
                       #INO_FB_Markers(IN_tNewMissionData := #TMP_tNewMisMark,
                                             IN_xStandardFBCall := FALSE,
                                             INO_xCallAddTank := #TMP_xCallAddTank,
                                             INO_tEnc := "DB_Encoder",INO_tRibbon := "DB_RibbonData");

                   END_IF;
               END_FOR;
           END_IF;
       END_IF;
   END_IF;

   //Manage received big telegram
   IF #FB_TRecvBig.DONE THEN

       //Check the packet telegram
       #TMP_dSerializePos := 0;
       #TMP_iReturn := Deserialize(SRC_ARRAY:=#AUX_rgb1000RecvBytePck, DEST_VARIABLE=>#TMP_dValue, POS:=#TMP_dSerializePos);

       IF #TMP_dValue = #DPLATEPACKTIDENT THEN

           #TMP_dSerializePos := 0;
           #TMP_iReturn := Deserialize(SRC_ARRAY:=#AUX_rgb1000RecvBytePck, DEST_VARIABLE=>#AUX_tPlatePacket, POS:=#TMP_dSerializePos);

           //Copy the plate to the buffer
           IF #AUX_dNumPlatePacket < #DMAXPLATEPACKET THEN

               #AUX_rgtPlatePacketArray[#AUX_dNumPlatePacket] := #AUX_tPlatePacket;
               #AUX_dNumPlatePacket+=1;

           END_IF;

       END_IF;
   END_IF;

   //Convert the plate data and make available for tracking
   IF #AUX_dNumPlatePacket > 0 AND #INO_tCaps.xInsertCapOnTrack = FALSE THEN

       #INO_tCaps.tNewCapToInsert := #INO_tCaps.tEmptyCap;

       #INO_tCaps.tNewCapToInsert.dID := #AUX_rgtPlatePacketArray[0].dCapID;
       #INO_tCaps.tNewCapToInsert.dHeadPositionBTC := #AUX_rgtPlatePacketArray[0].dPlateHead_cmm;
       #INO_tCaps.tNewCapToInsert.dTailPositionBTC := #AUX_rgtPlatePacketArray[0].dPlateHead_cmm + #AUX_rgtPlatePacketArray[0].dCapLength_cmm;


       #INO_tCaps.tNewCapToInsert.dLength_cmm := #AUX_rgtPlatePacketArray[0].dCapLength_cmm;

   //    IF "InsertStripe" THEN
   //        #INO_tCaps.tNewCapToInsert.dLength_cmm := 30000;//#AUX_rgtPlatePacketArray[0].dCapLength_cmm;
   //        #AUX_rgtPlatePacketArray[0].rgdDestMain[#TMP_dIndex] := "DCULLETDESTMASK";  
   //    "InsertStripe" := FALSE;
   //    END_IF;

    //   IF #AUX_rgtPlatePacketArray[0].rgdDestMain[0].%X1 OR #AUX_rgtPlatePacketArray[0].rgdDestMain[0].%X2 THEN
    //       #AUX_rgtPlatePacketArray[0].rgdDestMain[0] := "DCULLETDESTMASK";  
    //   
    //       
    //   END_IF;

   //                  #TMP_tNewMisMark.dMarkerID := 3;
   //                    #TMP_tNewMisMark.dMissionID := #AUX_rgtPlatePacketArray[0].dCapID;
   //                    #TMP_tNewMisMark.dPlateID := #AUX_rgtPlatePacketArray[0].rgdLiteID[0];
   //                    #TMP_tNewMisMark.dSpotSpace_cmm := 50;
   //                    #TMP_tNewMisMark.dXPosition_cmm := #AUX_rgtPlatePacketArray[0].dPlateHead_cmm;
   //                    #TMP_tNewMisMark.dYPosition_cmm := (#AUX_rgtPlatePacketArray[0].dTotCapWidth_cmm / -2) + #AUX_rgtPlatePacketArray[0].dWanderRec_cmm ;
   //                    #TMP_xCallAddTank := TRUE;
   //
   //                    #INO_FB_Markers(IN_tNewMissionData := #TMP_tNewMisMark,
   //                                          IN_xStandardFBCall := FALSE,
   //                                          INO_xCallAddTank := #TMP_xCallAddTank,
   //                                          INO_tEnc := "DB_Encoder",INO_tRibbon := "DB_RibbonData");

       #INO_tCaps.tNewCapToInsert.dWidth_cmm := #AUX_rgtPlatePacketArray[0].dTotCapWidth_cmm;
       #INO_tCaps.tNewCapToInsert.dThick_cmm := #AUX_rgtPlatePacketArray[0].dCapThick_cmm;
       #INO_tCaps.tNewCapToInsert.dIndex := #AUX_rgtPlatePacketArray[0].dIndexPlateConv;
       #INO_tCaps.tNewCapToInsert.dFormat := 0;
       #INO_tCaps.tNewCapToInsert.dNumLites := #AUX_rgtPlatePacketArray[0].dNumLiteCap;
       #INO_tCaps.tNewCapToInsert.dReqGapForConv_cmm := 0;
       #INO_tCaps.tNewCapToInsert.dMaxCapInConv := #AUX_rgtPlatePacketArray[0].dMaxPlateConv;
       #INO_tCaps.tNewCapToInsert.dConvTotLength_cmm := #AUX_rgtPlatePacketArray[0].dConvLength_cmm;
       #INO_tCaps.tNewCapToInsert.dMinWidth_cmm := #AUX_rgtPlatePacketArray[0].dMinWidth_cmm;
       #INO_tCaps.tNewCapToInsert.dMaxWidth_cmm := #AUX_rgtPlatePacketArray[0].dMaxWidth_cmm;
       #INO_tCaps.tNewCapToInsert.dGrossWidth_cmm := #INO_tOptimizer.tHMR.rgtRibbonData[#INO_tOptimizer.tHMW.dSelectRibbonDataSource].dGrossWidth_cmm;
       #INO_tCaps.tNewCapToInsert.dNetWidth_cmm := #INO_tOptimizer.tHMR.rgtRibbonData[#INO_tOptimizer.tHMW.dSelectRibbonDataSource].dNetWidth_cmm;
       #INO_tCaps.tNewCapToInsert.dDEdgeOpSide_cmm := #AUX_rgtPlatePacketArray[0].dTrimWidthOper_cmm;
       #INO_tCaps.tNewCapToInsert.dDEdgeOppOpSide_cmm := #AUX_rgtPlatePacketArray[0].dTrimWidthOpOper_cmm;
       #INO_tCaps.tNewCapToInsert.dTEdgeOpSide_cmm := #AUX_rgtPlatePacketArray[0].dTripleEdgeOpSide_cmm;
       #INO_tCaps.tNewCapToInsert.dTEdgeOppOpSide_cmm := #AUX_rgtPlatePacketArray[0].dTripleEdgeOppoOpSide_cmm;
       #INO_tCaps.tNewCapToInsert.dStartCutWander_cmm := #AUX_rgtPlatePacketArray[0].dWanderRec_cmm;
       #INO_tCaps.tNewCapToInsert.dEndCutWander_cmm := #AUX_rgtPlatePacketArray[0].dWanderRec_cmm;
       #INO_tCaps.tNewCapToInsert.dNetWander_cmm := #INO_tOptimizer.tHMR.rgtRibbonData[#INO_tOptimizer.tHMW.dSelectWanderDataSource].dNetWander_cmm;
       #INO_tCaps.tNewCapToInsert.dGrossWander_cmm := #INO_tOptimizer.tHMR.rgtRibbonData[#INO_tOptimizer.tHMW.dSelectWanderDataSource].dGrossWander_cmm;
       #INO_tCaps.tNewCapToInsert.dColor := #AUX_rgtPlatePacketArray[0].dColorID;
       #INO_tCaps.tNewCapToInsert.dFixedCapProductionID := #AUX_rgtPlatePacketArray[0].dFixedCapProdId;
       #INO_tCaps.tNewCapToInsert.tRequests.xYCutSampleTest := #AUX_rgtPlatePacketArray[0].tGeneralFlags.xYCutSampleTest;
       #INO_tCaps.tNewCapToInsert.tRequests.xIsCapFixed := #AUX_rgtPlatePacketArray[0].tGeneralFlags.xIsFixedCap;

       #INO_tCaps.tNewCapToInsert.strColorDescr := '';
       #INO_tCaps.tNewCapToInsert.dSystemMeasure := 0;

       IF #AUX_rgtPlatePacketArray[0].dYBridgeToCut = 1 THEN

           #INO_tCaps.tNewCapToInsert.tRequests.tYCutsData[0].rgdHeadsPositions := #AUX_rgtPlatePacketArray[0].rgYBridgePos_cmm;

           GATHER(IN:=#AUX_rgtPlatePacketArray[0].rgxYHeadMask,
                  OUT=>#TMP_dwMask);

           #TMP_wMask := DWORD_TO_WORD(#TMP_dwMask);     

           SCATTER(IN:=#TMP_wMask,
                   OUT=>#INO_tCaps.tNewCapToInsert.tRequests.tYCutsData[0].rgxHeadsRequest);

           IF (#TMP_wMask <> 0) THEN
               #INO_tCaps.tNewCapToInsert.tRequests.tYCutsData[0].xUseThisBridge := TRUE;
           END_IF;

       ELSIF #AUX_rgtPlatePacketArray[0].dYBridgeToCut = 2 THEN

           #INO_tCaps.tNewCapToInsert.tRequests.tYCutsData[1].rgdHeadsPositions := #AUX_rgtPlatePacketArray[0].rgYBridgePos_cmm;

           GATHER(IN:=#AUX_rgtPlatePacketArray[0].rgxYHeadMask,
                  OUT=>#TMP_dwMask);

           #TMP_wMask := DWORD_TO_WORD(#TMP_dwMask);     

           SCATTER(IN:=#TMP_wMask,
                   OUT=>#INO_tCaps.tNewCapToInsert.tRequests.tYCutsData[1].rgxHeadsRequest);

           IF (#TMP_wMask <> 0) THEN
               #INO_tCaps.tNewCapToInsert.tRequests.tYCutsData[1].xUseThisBridge := TRUE;
           END_IF;
       END_IF;

       FOR #TMP_dIndex := 0 TO #DMAXXCUT_IND DO

           #INO_tCaps.tNewCapToInsert.tRequests.rgxXCutReqHead[#TMP_dIndex] := #AUX_rgtPlatePacketArray[0].rgxCutMissionHead[#TMP_dIndex];
           #INO_tCaps.tNewCapToInsert.tRequests.rgxXCutReqTail[#TMP_dIndex] := #AUX_rgtPlatePacketArray[0].rgxCutMissionTail[#TMP_dIndex + 24];

       END_FOR;

       #INO_tCaps.tNewCapToInsert.tRequests.xOptSelvedgeSel := NOT #AUX_rgtPlatePacketArray[0].tGeneralFlags.xAutoTrim;
       #INO_tCaps.tNewCapToInsert.tRequests.xOptSplitBarSel := NOT #AUX_rgtPlatePacketArray[0].tGeneralFlags.xAutoSnap;
       #INO_tCaps.tNewCapToInsert.tRequests.xOptSepRollSel := NOT #AUX_rgtPlatePacketArray[0].tGeneralFlags.xAutoSep;
       #INO_tCaps.tNewCapToInsert.tRequests.dReqTrim3OpSide := #AUX_rgtPlatePacketArray[0].dTripleEdgeHeadOpSide;
       #INO_tCaps.tNewCapToInsert.tRequests.dReqTrim2OpSide := #AUX_rgtPlatePacketArray[0].dExtBordOp;
       #INO_tCaps.tNewCapToInsert.tRequests.dReqTrim1OpSide :=  #AUX_rgtPlatePacketArray[0].dIntBordOp;
       #INO_tCaps.tNewCapToInsert.tRequests.dReqTrim3OppOpSide := #AUX_rgtPlatePacketArray[0].dTripleEdgeHeadOppoOpSide;
       #INO_tCaps.tNewCapToInsert.tRequests.dReqTrim2OppOpSide := #AUX_rgtPlatePacketArray[0].dExtBordOppoOp;
       #INO_tCaps.tNewCapToInsert.tRequests.dReqTrim1OppOpSide := #AUX_rgtPlatePacketArray[0].dIntBordOp;
       #INO_tCaps.tNewCapToInsert.tRequests.rgdReqSplitBarSel := #AUX_rgtPlatePacketArray[0].rgdBumps;
       #INO_tCaps.tNewCapToInsert.tRequests.xIsCapFixed := #AUX_rgtPlatePacketArray[0].tGeneralFlags.xIsFixedCap;

       GATHER(IN:=#AUX_rgtPlatePacketArray[0].rgxChevrons,
              OUT=>#TMP_dwMask);

       #INO_tCaps.tNewCapToInsert.tRequests.rgbSeparatorSelect[3] := DWORD_TO_BYTE(SHR(IN:=#TMP_dwMask, N:=24));
       #INO_tCaps.tNewCapToInsert.tRequests.rgbSeparatorSelect[2] := DWORD_TO_BYTE(SHR(IN:=SHL(IN:=#TMP_dwMask,N:= 8), N:=24));
       #INO_tCaps.tNewCapToInsert.tRequests.rgbSeparatorSelect[1] := DWORD_TO_BYTE(SHR(IN:=SHL(IN:=#TMP_dwMask,N:= 16), N:=24));
       #INO_tCaps.tNewCapToInsert.tRequests.rgbSeparatorSelect[0] := DWORD_TO_BYTE(SHR(IN:=SHL(IN:=#TMP_dwMask,N:= 24), N:=24));

       #INO_tCaps.tNewCapToInsert.tRequests.xUpdateDataBPSA := TRUE;
       #INO_tCaps.tNewCapToInsert.tRequests.xUpdateDataBPSB := TRUE;
       #INO_tCaps.tNewCapToInsert.tRequests.xWandContinue := FALSE;

       FOR #TMP_dIndex := 0 TO #AUX_rgtPlatePacketArray[0].dNumLiteCap - 1 DO

           #INO_tCaps.tNewCapToInsert.rgtLites[#TMP_dIndex].dID := #AUX_rgtPlatePacketArray[0].rgdLiteID[#TMP_dIndex];
           #INO_tCaps.tNewCapToInsert.rgtLites[#TMP_dIndex].dProductionID := #AUX_rgtPlatePacketArray[0].rgdProductionID[#TMP_dIndex];
           #INO_tCaps.tNewCapToInsert.rgtLites[#TMP_dIndex].strProdDescr := '';
           #INO_tCaps.tNewCapToInsert.rgtLites[#TMP_dIndex].dQualityID := #AUX_rgtPlatePacketArray[0].rgdQualityID[#TMP_dIndex];
           #INO_tCaps.tNewCapToInsert.rgtLites[#TMP_dIndex].strQualityDescr := '';
           #INO_tCaps.tNewCapToInsert.rgtLites[#TMP_dIndex].dCameraRecipeID := #AUX_rgtPlatePacketArray[0].dGeomID;
           #INO_tCaps.tNewCapToInsert.rgtLites[#TMP_dIndex].dWidth_cmm := #AUX_rgtPlatePacketArray[0].rgdLiteWidth_cmm[#TMP_dIndex];
           #INO_tCaps.tNewCapToInsert.rgtLites[#TMP_dIndex].dBarycentre_cmm := 0;
           #INO_tCaps.tNewCapToInsert.rgtLites[#TMP_dIndex].dCulletCause := #AUX_rgtPlatePacketArray[0].rgdCulletCause[#TMP_dIndex];
           #INO_tCaps.tNewCapToInsert.rgtLites[#TMP_dIndex].rgxLayers[0] := #AUX_rgtPlatePacketArray[0].rgtLiteFlags[#TMP_dIndex].xPow1Req;
           #INO_tCaps.tNewCapToInsert.rgtLites[#TMP_dIndex].rgxLayers[1] := #AUX_rgtPlatePacketArray[0].rgtLiteFlags[#TMP_dIndex].xPow2Req;
           #INO_tCaps.tNewCapToInsert.rgtLites[#TMP_dIndex].dMainDestination := #AUX_rgtPlatePacketArray[0].rgdDestMain[#TMP_dIndex];
           #INO_tCaps.tNewCapToInsert.rgtLites[#TMP_dIndex].dAltDestination := #AUX_rgtPlatePacketArray[0].rgdDestAlt[#TMP_dIndex];
           #INO_tCaps.tNewCapToInsert.rgtLites[#TMP_dIndex].d2ndDestionation := #AUX_rgtPlatePacketArray[0].rgdDest2Nd[#TMP_dIndex];

           #INO_tCaps.tNewCapToInsert.rgtLites[#TMP_dIndex].dMainDestination := #AUX_rgtPlatePacketArray[0].rgdDestMain[#TMP_dIndex];
           #INO_tCaps.tNewCapToInsert.rgtLites[#TMP_dIndex].dAltDestination := #AUX_rgtPlatePacketArray[0].rgdDestAlt[#TMP_dIndex];
           #INO_tCaps.tNewCapToInsert.rgtLites[#TMP_dIndex].d2ndDestionation := #AUX_rgtPlatePacketArray[0].rgdDest2Nd[#TMP_dIndex];

           #INO_tCaps.tNewCapToInsert.rgtLites[#TMP_dIndex].tRequests.dMapLaserHeadOp := 0;
           #INO_tCaps.tNewCapToInsert.rgtLites[#TMP_dIndex].tRequests.dMapLaserHeadOppOp := 0;
           #INO_tCaps.tNewCapToInsert.rgtLites[#TMP_dIndex].xSaturationPlate := #AUX_rgtPlatePacketArray[0].rgtLiteFlags[#TMP_dIndex].xSatPlate;
           #INO_tCaps.tNewCapToInsert.rgtLites[#TMP_dIndex].tRequests.xGeomInsp := #AUX_rgtPlatePacketArray[0].rgtLiteFlags[#TMP_dIndex].xGeomInsp;

       END_FOR;

       #AUX_dNumPlatePacket-= 1;

       IF #AUX_dNumPlatePacket > 0 THEN
           #TMP_iReturn := MOVE_BLK_VARIANT(SRC:=#AUX_rgtPlatePacketArray, COUNT:=DINT_TO_UDINT(#AUX_dNumPlatePacket), SRC_INDEX:=1, DEST_INDEX:=0, DEST=>#AUX_rgtPlatePacketArray);
       END_IF;

       #INO_tCaps.xInsertCapOnTrack := TRUE;

   END_IF;
END_FUNCTION_BLOCK

// folder: 03_Programs_Logics/MCC1200/06_InitUtility

FUNCTION_BLOCK "GP_OB_Initialize"   // FB7, SCL
TITLE = OB Service flags
{ S7_Optimized_Access := 'TRUE' }
AUTHOR : Cigliutt
FAMILY : GP
VERSION : 1.1
// This FB will provide the following information: 1# OB duration time 2# Timer clock and OS. IMPORTANT!!! This FB must be initialized each OB100 call, and must be called for each OB!
   VAR_INPUT
      IN_xInitialize : Bool;   // Initialize values (OB100 call)
   END_VAR
   VAR
      STC_rlLastExecValue_s : LReal;   // Last execution tick value [s]
      STC_rlReminder_s : Real;   // Reminder from last execution [ms]
      STC_dElapsed_100ms_ms : DInt;   // Elapsed time for 0.1s
      STC_dElapsed_200ms_ms : DInt;   // Elapsed time for 0.2s
      STC_dElapsed_400ms_ms : DInt;   // Elapsed time for 0.4s
      STC_dElapsed_500ms_ms : DInt;   // Elapsed time for 0.5s
      STC_dElapsed_800ms_ms : DInt;   // Elapsed time for 0.8s
      STC_dElapsed_1s_ms : DInt;   // Elapsed time for 1s
      STC_dElapsed_2s_ms : DInt;   // Elapsed time for 2s
      STC_dElapsed_5s_ms : DInt;   // Elapsed time for 5s
      STC_dElapsed_10s_ms : DInt;   // Elapsed time for 10s
      STC_dElapsed_30s_ms : DInt;   // Elapsed time for 30s
      STC_dElapsed_1min_ms : DInt;   // Elapsed time for 1min
      STC_dElapsed_2min_ms : DInt;   // Elapsed time for 2min
      STC_dElapsed_10min_ms : DInt;   // Elapsed time for 10min
      STC_dElapsed_30min_ms : DInt;   // Elapsed time for 30min
      STC_dElapsed_1h_ms : DInt;   // Elapsed time for 1h
      OUT_dExecutionTime_ms : DInt;   // OB Execution time [ms]
      OUT_dMinExecutionTime_ms : DInt;   // OB Maximum execution time [ms]
      OUT_dMaxExecutionTime_ms : DInt;   // OB Minimum execution time [ms]
      OUT_xOs_100ms : Bool;   // OS each 100ms
      OUT_xOs_200ms : Bool;   // OS each 200ms
      OUT_xOs_400ms : Bool;   // OS each 400ms
      OUT_xOs_500ms : Bool;   // OS each 500ms
      OUT_xOs_800ms : Bool;   // OS each 800ms
      OUT_xOs_1s : Bool;   // OS each 1s
      OUT_xOs_2s : Bool;   // OS each 2s
      OUT_xOs_5s : Bool;   // OS each 5s
      OUT_xOs_10s : Bool;   // OS each 10s
      OUT_xOs_30s : Bool;   // OS each 30s
      OUT_xOs_1min : Bool;   // OS each 1min
      OUT_xOs_2min : Bool;   // OS each 2min
      OUT_xOs_10min : Bool;   // OS each 10min
      OUT_xOs_30min : Bool;   // OS each 30min
      OUT_xOs_1h : Bool;   // OS each 1h
      OUT_xClock_100ms : Bool;   // Clock 100ms
      OUT_xClock_200ms : Bool;   // Clock 200ms
      OUT_xClock_400ms : Bool;   // Clock 400ms
      OUT_xClock_500ms : Bool;   // Clock 500ms
      OUT_xClock_800ms : Bool;   // Clock 800ms
      OUT_xClock_1s : Bool;   // Clock 1s
      OUT_xClock_2s : Bool;   // Clock 2s
      OUT_xClock_5s : Bool;   // Clock 5s
      OUT_xClock_10s : Bool;   // Clock 10s
      OUT_xClock_30s : Bool;   // Clock 30s
      OUT_xClock_1min : Bool;   // Clock 1min
      OUT_xClock_2min : Bool;   // Clock 2min
      OUT_xClock_10min : Bool;   // Clock 10min
      OUT_xClock_30min : Bool;   // Clock 30min
      OUT_xClock_1h : Bool;   // Clock 1h
      OUT_xDebugOFF : Bool;   // Commisioning bit - Always OFF
      OUT_xDebugON : Bool;   // Commisioning bit - Always ON
   END_VAR
   VAR_TEMP
      TMP_rlActualExecutionTime : Real;   // ActualExecutionTime [ms]
      TMP_rlActualExecutionTimeRound : Real;   // Rounded execution time [ms]
      TMP_rlActualExecutionTimeCalculated : Real;
   END_VAR
   VAR CONSTANT
      CONST_DTICK_100MS : DInt := 100;
      CONST_DTICK_200MS : DInt := 200;
      CONST_DTICK_400MS : DInt := 400;
      CONST_DTICK_500MS : DInt := 500;
      CONST_DTICK_800MS : DInt := 800;
      CONST_DTICK_1S : DInt := 1000;
      CONST_DTICK_2S : DInt := 2000;
      CONST_DTICK_5S : DInt := 5000;
      CONST_DTICK_10S : DInt := 10000;
      CONST_DTICK_30S : DInt := 30000;
      CONST_DTICK_1MIN : DInt := 60000;
      CONST_DTICK_2MIN : DInt := 120000;
      CONST_DTICK_10MIN : DInt := 600000;
      CONST_DTICK_30MIN : DInt := 1800000;
      CONST_DTICK_1H : DInt := 86400000;
      CONST_DMAX_INT : DInt := 16#7FFF_FFFF;
   END_VAR
BEGIN
   //Initialize OS bits
   #OUT_xOs_100ms := false;
   #OUT_xOs_200ms := false;
   #OUT_xOs_400ms := false;
   #OUT_xOs_500ms := false;
   #OUT_xOs_800ms := false;
   #OUT_xOs_1s := false;
   #OUT_xOs_2s := false;
   #OUT_xOs_5s := false;
   #OUT_xOs_10s := false;
   #OUT_xOs_30s := false;
   #OUT_xOs_1min := false;
   #OUT_xOs_2min := false;
   #OUT_xOs_10min := false;
   #OUT_xOs_30min := false;
   #OUT_xOs_1h := false;

   //Initialize FB execution
   IF #IN_xInitialize = true THEN


       #IN_xInitialize := false;

       #OUT_dExecutionTime_ms := 0;
       #OUT_dMinExecutionTime_ms := #CONST_DMAX_INT;
       #OUT_dMaxExecutionTime_ms := 0;
       #OUT_xClock_100ms := false;
       #OUT_xClock_200ms := false;
       #OUT_xClock_400ms := false;
       #OUT_xClock_500ms := false;
       #OUT_xClock_800ms := false;
       #OUT_xClock_1s := false;
       #OUT_xClock_2s := false;
       #OUT_xClock_5s := false;
       #OUT_xClock_10s := false;
       #OUT_xClock_30s := false;
       #OUT_xClock_1min := false;
       #OUT_xClock_2min := false;
       #OUT_xClock_10min := false;
       #OUT_xClock_30min := false;
       #OUT_xClock_1h := false;

       #STC_dElapsed_100ms_ms := 0;
       #STC_dElapsed_200ms_ms := 0;
       #STC_dElapsed_400ms_ms := 0;
       #STC_dElapsed_500ms_ms := 0;
       #STC_dElapsed_800ms_ms := 0;
       #STC_dElapsed_1s_ms := 0;
       #STC_dElapsed_2s_ms := 0;
       #STC_dElapsed_5s_ms := 0;
       #STC_dElapsed_10s_ms := 0;
       #STC_dElapsed_30s_ms := 0;
       #STC_dElapsed_1min_ms := 0;
       #STC_dElapsed_2min_ms := 0;
       #STC_dElapsed_10min_ms := 0;
       #STC_dElapsed_30min_ms := 0;
       #STC_dElapsed_1h_ms := 0;
       #STC_rlLastExecValue_s := 0;
       #STC_rlReminder_s := 0;
       #STC_rlLastExecValue_s := 0;

   END_IF;
   //***** CALCULATE OB EXECUTION TIME ***** 
   //Take the execution time from the CPU
   #TMP_rlActualExecutionTime := LREAL_TO_REAL(RUNTIME(MEM := #STC_rlLastExecValue_s));

   //Convert from [s] to [ms]
   #TMP_rlActualExecutionTime := #TMP_rlActualExecutionTime * 1000.0;

   //Add the reminder of the last cycle
   #TMP_rlActualExecutionTimeCalculated := #TMP_rlActualExecutionTime + #STC_rlReminder_s;
   //Calculate the rounded value
   #TMP_rlActualExecutionTimeRound := ROUND_REAL(#TMP_rlActualExecutionTimeCalculated);
   #OUT_dExecutionTime_ms := ROUND_DINT(#TMP_rlActualExecutionTimeCalculated);

   //Save the reminder for the next cycle
   #STC_rlReminder_s := #TMP_rlActualExecutionTimeCalculated - #TMP_rlActualExecutionTimeRound;

   //Save the maximum scan value
   IF #OUT_dExecutionTime_ms > #OUT_dMaxExecutionTime_ms THEN
       #OUT_dMaxExecutionTime_ms := #OUT_dExecutionTime_ms;
   END_IF;

   //Save the minimum scan value
   IF #OUT_dExecutionTime_ms < #OUT_dMinExecutionTime_ms THEN
       #OUT_dMinExecutionTime_ms := #OUT_dExecutionTime_ms;
   END_IF;

   //***** CALCULATE SERVICES CLOCK *****

   //Increment counters for each clock
   #STC_dElapsed_100ms_ms := #STC_dElapsed_100ms_ms + #OUT_dExecutionTime_ms;
   #STC_dElapsed_200ms_ms := #STC_dElapsed_200ms_ms + #OUT_dExecutionTime_ms;
   #STC_dElapsed_400ms_ms := #STC_dElapsed_400ms_ms + #OUT_dExecutionTime_ms;
   #STC_dElapsed_500ms_ms := #STC_dElapsed_500ms_ms + #OUT_dExecutionTime_ms;
   #STC_dElapsed_800ms_ms := #STC_dElapsed_800ms_ms + #OUT_dExecutionTime_ms;
   #STC_dElapsed_1s_ms := #STC_dElapsed_1s_ms + #OUT_dExecutionTime_ms;
   #STC_dElapsed_2s_ms := #STC_dElapsed_2s_ms + #OUT_dExecutionTime_ms;
   #STC_dElapsed_5s_ms := #STC_dElapsed_5s_ms + #OUT_dExecutionTime_ms;
   #STC_dElapsed_10s_ms := #STC_dElapsed_10s_ms + #OUT_dExecutionTime_ms;
   #STC_dElapsed_30s_ms := #STC_dElapsed_30s_ms + #OUT_dExecutionTime_ms;
   #STC_dElapsed_1min_ms := #STC_dElapsed_1min_ms + #OUT_dExecutionTime_ms;
   #STC_dElapsed_2min_ms := #STC_dElapsed_2min_ms + #OUT_dExecutionTime_ms;
   #STC_dElapsed_10min_ms := #STC_dElapsed_10min_ms + #OUT_dExecutionTime_ms;
   #STC_dElapsed_30min_ms := #STC_dElapsed_30min_ms + #OUT_dExecutionTime_ms;
   #STC_dElapsed_1h_ms := #STC_dElapsed_1h_ms + #OUT_dExecutionTime_ms;

   //Calculate the 100ms
   IF #STC_dElapsed_100ms_ms >= #CONST_DTICK_100MS THEN
       #STC_dElapsed_100ms_ms := #STC_dElapsed_100ms_ms - #CONST_DTICK_100MS;

       #OUT_xOs_100ms := true;

       IF (#OUT_xClock_100ms = false) THEN
           #OUT_xClock_100ms := true;
       ELSE
           #OUT_xClock_100ms := false;
       END_IF;
   END_IF;

   //Calculate the 200ms
   IF #STC_dElapsed_200ms_ms >= #CONST_DTICK_200MS THEN
       #STC_dElapsed_200ms_ms := #STC_dElapsed_200ms_ms - #CONST_DTICK_200MS;

       #OUT_xOs_200ms := true;

       IF (#OUT_xClock_200ms = false) THEN
           #OUT_xClock_200ms := true;
       ELSE
           #OUT_xClock_200ms := false;
       END_IF;
   END_IF;

   //Calculate the 400ms
   IF #STC_dElapsed_400ms_ms >= #CONST_DTICK_400MS THEN
       #STC_dElapsed_400ms_ms := #STC_dElapsed_400ms_ms - #CONST_DTICK_400MS;

       #OUT_xOs_400ms := true;

       IF (#OUT_xClock_400ms = false) THEN
           #OUT_xClock_400ms := true;
       ELSE
           #OUT_xClock_400ms := false;
       END_IF;
   END_IF;

   //Calculate the 500ms
   IF #STC_dElapsed_500ms_ms >= #CONST_DTICK_500MS THEN
       #STC_dElapsed_500ms_ms := #STC_dElapsed_500ms_ms - #CONST_DTICK_500MS;

       #OUT_xOs_500ms := true;

       IF (#OUT_xClock_500ms = false) THEN
           #OUT_xClock_500ms := true;
       ELSE
           #OUT_xClock_500ms := false;
       END_IF;
   END_IF;

   //Calculate the 800ms
   IF #STC_dElapsed_800ms_ms >= #CONST_DTICK_800MS THEN
       #STC_dElapsed_800ms_ms := #STC_dElapsed_800ms_ms - #CONST_DTICK_800MS;

       #OUT_xOs_800ms := true;

       IF (#OUT_xClock_800ms = false) THEN
           #OUT_xClock_800ms := true;
       ELSE
           #OUT_xClock_800ms := false;
       END_IF;
   END_IF;

   //Calculate the 1s
   IF #STC_dElapsed_1s_ms >= #CONST_DTICK_1S THEN
       #STC_dElapsed_1s_ms := #STC_dElapsed_1s_ms - #CONST_DTICK_1S;

       #OUT_xOs_1s := true;

       IF (#OUT_xClock_1s = false) THEN
           #OUT_xClock_1s := true;
       ELSE
           #OUT_xClock_1s := false;
       END_IF;
   END_IF;

   //Calculate the 2s
   IF #STC_dElapsed_2s_ms >= #CONST_DTICK_2S THEN
       #STC_dElapsed_2s_ms := #STC_dElapsed_2s_ms - #CONST_DTICK_2S;

       #OUT_xOs_2s := true;

       IF (#OUT_xClock_2s = false) THEN
           #OUT_xClock_2s := true;
       ELSE
           #OUT_xClock_2s := false;
       END_IF;
   END_IF;

   //Calculate the 5s
   IF #STC_dElapsed_5s_ms >= #CONST_DTICK_5S THEN
       #STC_dElapsed_5s_ms := #STC_dElapsed_5s_ms - #CONST_DTICK_5S;

       #OUT_xOs_5s := true;

       IF (#OUT_xClock_5s = false) THEN
           #OUT_xClock_5s := true;
       ELSE
           #OUT_xClock_5s := false;
       END_IF;
   END_IF;

   //Calculate the 10s
   IF #STC_dElapsed_10s_ms >= #CONST_DTICK_10S THEN
       #STC_dElapsed_10s_ms := #STC_dElapsed_10s_ms - #CONST_DTICK_10S;

       #OUT_xOs_10s := true;

       IF (#OUT_xClock_10s = false) THEN
           #OUT_xClock_10s := true;
       ELSE
           #OUT_xClock_10s := false;
       END_IF;
   END_IF;

   //Calculate the 30s
   IF #STC_dElapsed_30s_ms >= #CONST_DTICK_30S THEN
       #STC_dElapsed_30s_ms := #STC_dElapsed_30s_ms - #CONST_DTICK_30S;

       #OUT_xOs_30s := true;

       IF (#OUT_xClock_30s = false) THEN
           #OUT_xClock_30s := true;
       ELSE
           #OUT_xClock_30s := false;
       END_IF;
   END_IF;

   //Calculate the 1min
   IF #STC_dElapsed_1min_ms >= #CONST_DTICK_1MIN THEN
       #STC_dElapsed_1min_ms := #STC_dElapsed_1min_ms - #CONST_DTICK_1MIN;

       #OUT_xOs_1min := true;

       IF (#OUT_xClock_1min = false) THEN
           #OUT_xClock_1min := true;
       ELSE
           #OUT_xClock_1min := false;
       END_IF;
   END_IF;

   //Calculate the 2min
   IF #STC_dElapsed_2min_ms >= #CONST_DTICK_2MIN THEN
       #STC_dElapsed_2min_ms := #STC_dElapsed_2min_ms - #CONST_DTICK_2MIN;

       #OUT_xOs_2min := true;

       IF (#OUT_xClock_2min = false) THEN
           #OUT_xClock_2min := true;
       ELSE
           #OUT_xClock_2min := false;
       END_IF;
   END_IF;

   //Calculate the 10min
   IF #STC_dElapsed_10min_ms >= #CONST_DTICK_10MIN THEN
       #STC_dElapsed_10min_ms := #STC_dElapsed_10min_ms - #CONST_DTICK_10MIN;

       #OUT_xOs_10min := true;

       IF (#OUT_xClock_10min = false) THEN
           #OUT_xClock_10min := true;
       ELSE
           #OUT_xClock_10min := false;
       END_IF;
   END_IF;

   //Calculate the 30min
   IF #STC_dElapsed_30min_ms >= #CONST_DTICK_30MIN THEN
       #STC_dElapsed_30min_ms := #STC_dElapsed_30min_ms - #CONST_DTICK_30MIN;

       #OUT_xOs_30min := true;

       IF (#OUT_xClock_30min = false) THEN
           #OUT_xClock_30min := true;
       ELSE
           #OUT_xClock_30min := false;
       END_IF;
   END_IF;

   //Calculate the 1h
   IF #STC_dElapsed_1h_ms >= #CONST_DTICK_1H THEN
       #STC_dElapsed_1h_ms := #STC_dElapsed_1h_ms - #CONST_DTICK_1H;

       #OUT_xOs_1h := true;

       IF (#OUT_xClock_1h = false) THEN
           #OUT_xClock_1h := true;
       ELSE
           #OUT_xClock_1h := false;
       END_IF;
   END_IF;
END_FUNCTION_BLOCK

// folder: 03_Programs_Logics/MCC1200/09_Zone

FUNCTION "Z200_Faults" : Void   // FC1, LAD
{ S7_Optimized_Access := 'TRUE' }
VERSION : 0.1
   VAR_TEMP
      TMP_dwValue : DWord;
   END_VAR
BEGIN

REGION Network 1 (SCL): Reset alarms
   IF "Z201".tmOFF_ResetAlarm.OUT_xDone OR "ZUPS".tmOFF_ResetAlarm.OUT_xDone THEN

       #TMP_dwValue := 0;

       SCATTER(IN:=#TMP_dwValue,
               OUT=>"DB_Z200_HMI".tALM.tE);

       SCATTER(IN:=#TMP_dwValue,
               OUT=>"DB_Z200_HMI".tALM.tS);

       SCATTER(IN:=#TMP_dwValue,
               OUT=>"DB_Z200_HMI".tALM.tF);

       SCATTER(IN:=#TMP_dwValue,
               OUT=>"DB_Z200_HMI".tALM.tW);

   END_IF;
END_REGION

REGION Network 2: ### STOPPING FAULTS ###
END_REGION

REGION Network 3: Anomalies / ### FAULTS ###
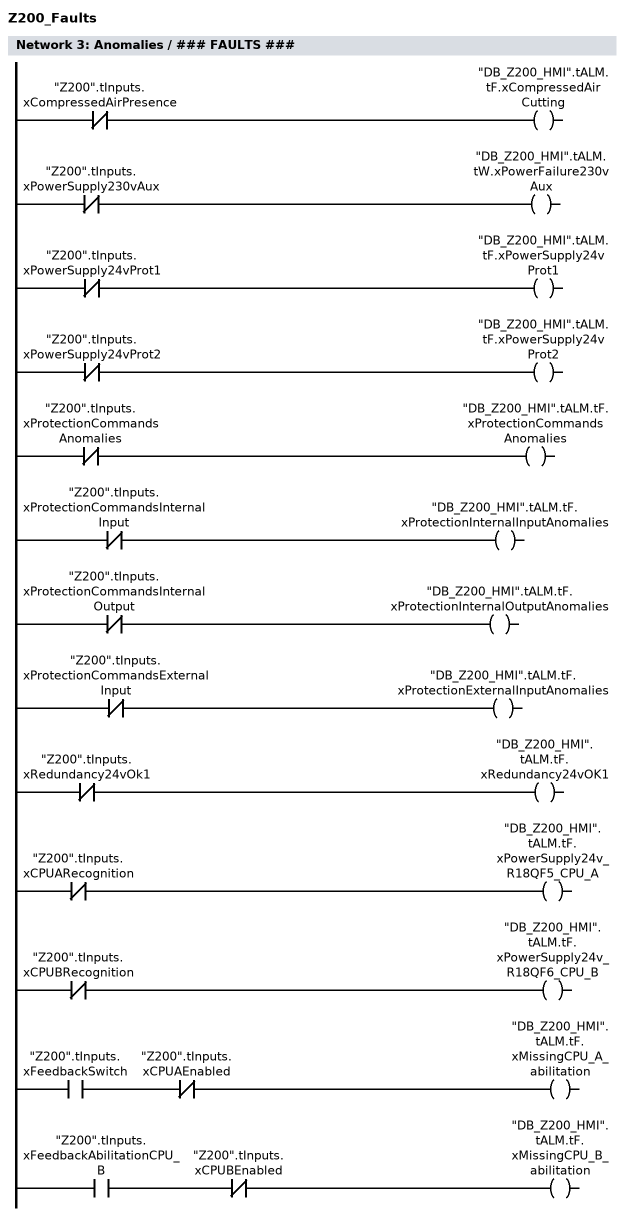
   RUNG wire#powerrail
      I_Contact( "Z200".tInputs.xCompressedAirPresence )
      Coil( "DB_Z200_HMI".tALM.tF.xCompressedAirCutting )
   END_RUNG
   RUNG wire#powerrail
      I_Contact( "Z200".tInputs.xPowerSupply230vAux )
      Coil( "DB_Z200_HMI".tALM.tW.xPowerFailure230vAux )
   END_RUNG
   RUNG wire#powerrail
      I_Contact( "Z200".tInputs.xPowerSupply24vProt1 )
      Coil( "DB_Z200_HMI".tALM.tF.xPowerSupply24vProt1 )
   END_RUNG
   RUNG wire#powerrail
      I_Contact( "Z200".tInputs.xPowerSupply24vProt2 )
      Coil( "DB_Z200_HMI".tALM.tF.xPowerSupply24vProt2 )
   END_RUNG
   RUNG wire#powerrail
      I_Contact( "Z200".tInputs.xProtectionCommandsAnomalies )
      Coil( "DB_Z200_HMI".tALM.tF.xProtectionCommandsAnomalies )
   END_RUNG
   RUNG wire#powerrail
      I_Contact( "Z200".tInputs.xProtectionCommandsInternalInput )
      Coil( "DB_Z200_HMI".tALM.tF.xProtectionInternalInputAnomalies )
   END_RUNG
   RUNG wire#powerrail
      I_Contact( "Z200".tInputs.xProtectionCommandsInternalOutput )
      Coil( "DB_Z200_HMI".tALM.tF.xProtectionInternalOutputAnomalies )
   END_RUNG
   RUNG wire#powerrail
      I_Contact( "Z200".tInputs.xProtectionCommandsExternalInput )
      Coil( "DB_Z200_HMI".tALM.tF.xProtectionExternalInputAnomalies )
   END_RUNG
   RUNG wire#powerrail
      I_Contact( "Z200".tInputs.xRedundancy24vOk1 )
      Coil( "DB_Z200_HMI".tALM.tF.xRedundancy24vOK1 )
   END_RUNG
   RUNG wire#powerrail
      I_Contact( "Z200".tInputs.xCPUARecognition )
      Coil( "DB_Z200_HMI".tALM.tF.xPowerSupply24v_R18QF5_CPU_A )
   END_RUNG
   RUNG wire#powerrail
      I_Contact( "Z200".tInputs.xCPUBRecognition )
      Coil( "DB_Z200_HMI".tALM.tF.xPowerSupply24v_R18QF6_CPU_B )
   END_RUNG
   RUNG wire#powerrail
      Contact( "Z200".tInputs.xFeedbackSwitch )
      I_Contact( "Z200".tInputs.xCPUAEnabled )
      Coil( "DB_Z200_HMI".tALM.tF.xMissingCPU_A_abilitation )
   END_RUNG
   RUNG wire#powerrail
      Contact( "Z200".tInputs.xFeedbackAbilitationCPU_B )
      I_Contact( "Z200".tInputs.xCPUBEnabled )
      Coil( "DB_Z200_HMI".tALM.tF.xMissingCPU_B_abilitation )
   END_RUNG
   // the same network as SCL:
   "DB_Z200_HMI".tALM.tF.xCompressedAirCutting := NOT "Z200".tInputs.xCompressedAirPresence;
   "DB_Z200_HMI".tALM.tW.xPowerFailure230vAux := NOT "Z200".tInputs.xPowerSupply230vAux;
   "DB_Z200_HMI".tALM.tF.xPowerSupply24vProt1 := NOT "Z200".tInputs.xPowerSupply24vProt1;
   "DB_Z200_HMI".tALM.tF.xPowerSupply24vProt2 := NOT "Z200".tInputs.xPowerSupply24vProt2;
   "DB_Z200_HMI".tALM.tF.xProtectionCommandsAnomalies := NOT "Z200".tInputs.xProtectionCommandsAnomalies;
   "DB_Z200_HMI".tALM.tF.xProtectionInternalInputAnomalies := NOT "Z200".tInputs.xProtectionCommandsInternalInput;
   "DB_Z200_HMI".tALM.tF.xProtectionInternalOutputAnomalies := NOT "Z200".tInputs.xProtectionCommandsInternalOutput;
   "DB_Z200_HMI".tALM.tF.xProtectionExternalInputAnomalies := NOT "Z200".tInputs.xProtectionCommandsExternalInput;
   "DB_Z200_HMI".tALM.tF.xRedundancy24vOK1 := NOT "Z200".tInputs.xRedundancy24vOk1;
   "DB_Z200_HMI".tALM.tF.xPowerSupply24v_R18QF5_CPU_A := NOT "Z200".tInputs.xCPUARecognition;
   "DB_Z200_HMI".tALM.tF.xPowerSupply24v_R18QF6_CPU_B := NOT "Z200".tInputs.xCPUBRecognition;
   "DB_Z200_HMI".tALM.tF.xMissingCPU_A_abilitation := "Z200".tInputs.xFeedbackSwitch AND NOT "Z200".tInputs.xCPUAEnabled;
   "DB_Z200_HMI".tALM.tF.xMissingCPU_B_abilitation := "Z200".tInputs.xFeedbackAbilitationCPU_B AND NOT "Z200".tInputs.xCPUBEnabled;
END_REGION

REGION Network 4 (SCL): Calculate comulative status
   GATHER(IN:="DB_Z200_HMI".tALM.tE,
              OUT=>#TMP_dwValue);


       GATHER(IN:="DB_Z200_HMI".tALM.tS,
              OUT=>#TMP_dwValue);

   IF #TMP_dwValue <> 0 THEN
       "Z200".ST_xZoneStoppingFaults := TRUE;
   ELSE
       "Z200".ST_xZoneStoppingFaults := FALSE;
   END_IF;

   GATHER(IN:="DB_Z200_HMI".tALM.tF,
              OUT=>#TMP_dwValue);

   IF #TMP_dwValue <> 0 THEN
       "Z200".ST_xZoneFaults := TRUE;
   ELSE
       "Z200".ST_xZoneFaults := FALSE;
   END_IF;

   GATHER(IN:="DB_Z200_HMI".tALM.tW,
              OUT=>#TMP_dwValue);

   IF #TMP_dwValue <> 0 THEN
       "Z200".ST_xZoneWarnings := TRUE;
   ELSE
       "Z200".ST_xZoneWarnings := FALSE;
   END_IF;

   IF "Z200".ST_xZoneStoppingFaults AND"Z200".ST_xZoneFaults THEN
       "Z200".ST_xZoneError := TRUE;
   ELSE
       "Z200".ST_xZoneError := FALSE;
   END_IF;
END_REGION
END_FUNCTION

FUNCTION "Z200_Logics" : Void   // FC7, LAD
{ S7_Optimized_Access := 'TRUE' }
VERSION : 0.1
   VAR_TEMP
      TMP_xGeneralMcc : Bool;
      TMP_xLocalMcc : Bool;
      TMP_rlVal : LReal;
   END_VAR
BEGIN

REGION Network 1: #### CONSTANTS ####
END_REGION

REGION Network 2 (SCL): ### SIMULATION ###
   IF "SIMULATION_ACTIVE" THEN

       "Z200".tInputs.xCPUAEnabled := TRUE;
       "Z200".tInputs.xCPUBEnabled := FALSE;
       "Z200".tInputs.xCPUARecognition := TRUE;
       "Z200".tInputs.xCPUBRecognition := FALSE;

       "Z200".tInputs.xCompressedAirPresence := TRUE;
       "Z200".tInputs.xProtectionCommandsAnomalies := TRUE;
       "Z200".tInputs.xProtectionCommandsInternalInput := TRUE;
       "Z200".tInputs.xProtectionCommandsInternalOutput := TRUE;
       "Z200".tInputs.xProtectionCommandsExternalInput := TRUE;
       "Z200".tInputs.xPowerSupply230vAux := TRUE;
       "Z200".tInputs.xRedundancy24vOk1 := TRUE;



       "Z200".tInputs.xMainEmergencyON := TRUE;
   END_IF;
   "TestTag64" := 0;
   "TestTag64".%X40 := 1;
END_REGION

REGION Network 3: #### MATCH ####
END_REGION

REGION Network 4: #### PLC ACTIVE ####
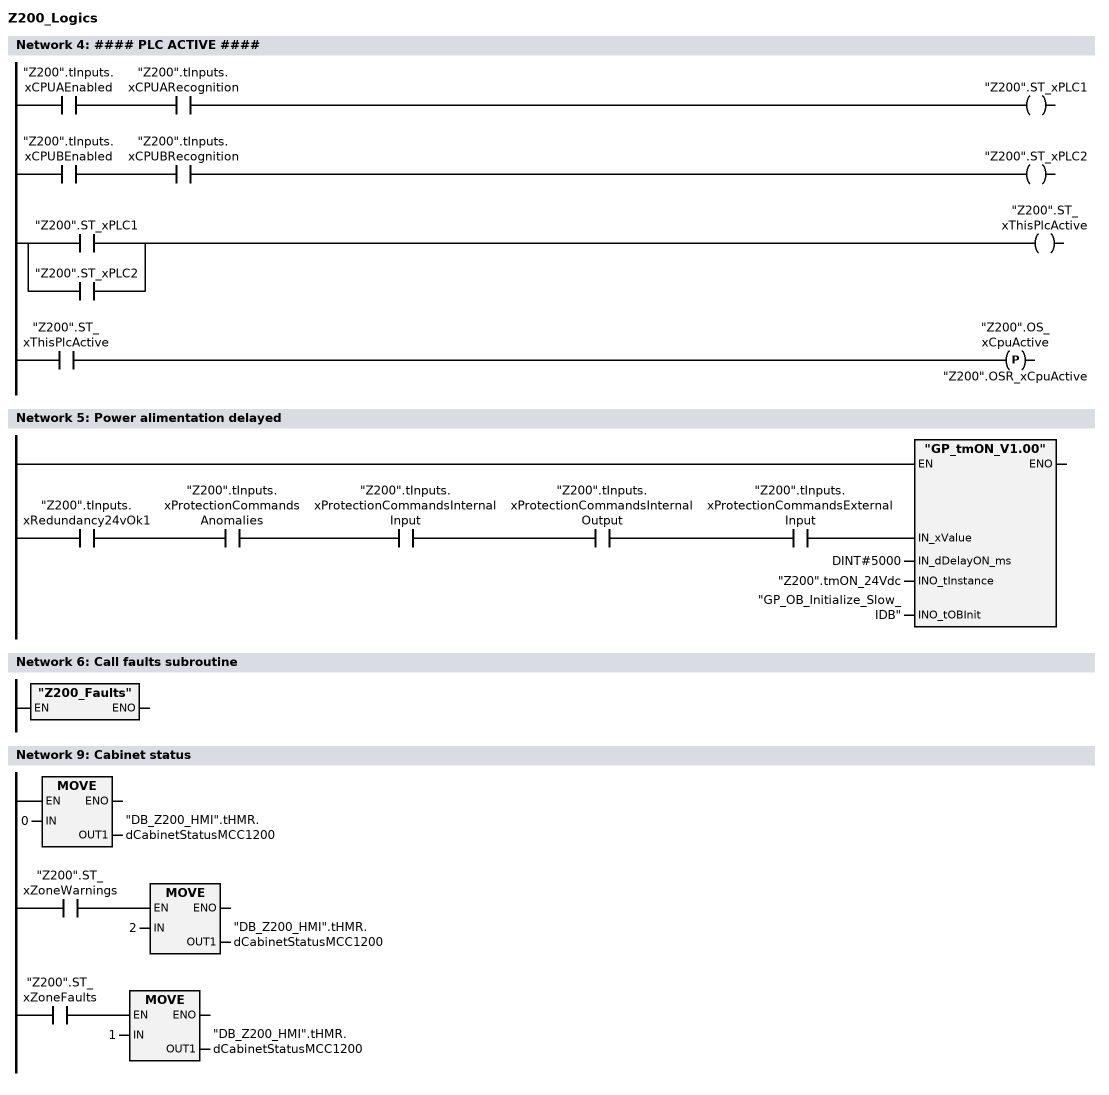
   "Z200".ST_xPLC1 := "Z200".tInputs.xCPUAEnabled AND "Z200".tInputs.xCPUARecognition;
   "Z200".ST_xPLC2 := "Z200".tInputs.xCPUBEnabled AND "Z200".tInputs.xCPUBRecognition;
   "Z200".ST_xThisPlcActive := "Z200".ST_xPLC1 OR "Z200".ST_xPLC2;
   "Z200".OS_xCpuActive := "Z200".ST_xThisPlcActive AND NOT "Z200".OSR_xCpuActive;   // rising edge
   "Z200".OSR_xCpuActive := "Z200".ST_xThisPlcActive;
END_REGION

REGION Network 5: Power alimentation delayed
   RUNG wire#powerrail
      "GP_tmON_V1.00"(IN_xValue := wire#w1, IN_dDelayON_ms := DINT#5000, INO_tInstance := "Z200".tmON_24Vdc, INO_tOBInit := "GP_OB_Initialize_Slow_IDB")
   END_RUNG
   RUNG wire#powerrail
      Contact( "Z200".tInputs.xRedundancy24vOk1 )
      Contact( "Z200".tInputs.xProtectionCommandsAnomalies )
      Contact( "Z200".tInputs.xProtectionCommandsInternalInput )
      Contact( "Z200".tInputs.xProtectionCommandsInternalOutput )
      Contact( "Z200".tInputs.xProtectionCommandsExternalInput )
   END_RUNG wire#w1
   // the same network as SCL:
   "GP_tmON_V1.00"(IN_xValue := "Z200".tInputs.xRedundancy24vOk1 AND "Z200".tInputs.xProtectionCommandsAnomalies AND "Z200".tInputs.xProtectionCommandsInternalInput AND "Z200".tInputs.xProtectionCommandsInternalOutput AND "Z200".tInputs.xProtectionCommandsExternalInput,
                   IN_dDelayON_ms := DINT#5000,
                   INO_tInstance := "Z200".tmON_24Vdc,
                   INO_tOBInit := "GP_OB_Initialize_Slow_IDB");
END_REGION

REGION Network 6: Call faults subroutine
   RUNG wire#powerrail
      "Z200_Faults"()
   END_RUNG
   // the same network as SCL:
   "Z200_Faults"();
END_REGION

REGION Network 7: #### START/STOP ZONE ####
END_REGION

REGION Network 8: #### HMI STATUSES ####
END_REGION

REGION Network 9: Cabinet status
   RUNG wire#powerrail
      Move(in := 0, out1 => "DB_Z200_HMI".tHMR.dCabinetStatusMCC1200)
   END_RUNG
   RUNG wire#powerrail
      Contact( "Z200".ST_xZoneWarnings )
      Move(in := 2, out1 => "DB_Z200_HMI".tHMR.dCabinetStatusMCC1200)
   END_RUNG
   RUNG wire#powerrail
      Contact( "Z200".ST_xZoneFaults )
      Move(in := 1, out1 => "DB_Z200_HMI".tHMR.dCabinetStatusMCC1200)
   END_RUNG
   // the same network as SCL:
   "DB_Z200_HMI".tHMR.dCabinetStatusMCC1200 := 0;
   IF "Z200".ST_xZoneWarnings THEN "DB_Z200_HMI".tHMR.dCabinetStatusMCC1200 := 2; END_IF;
   IF "Z200".ST_xZoneFaults THEN "DB_Z200_HMI".tHMR.dCabinetStatusMCC1200 := 1; END_IF;
END_REGION
END_FUNCTION

FUNCTION "Z200_Output" : Void   // FC14, LAD
{ S7_Optimized_Access := 'TRUE' }
VERSION : 0.1
   VAR CONSTANT
      CONST_DBREAKDOWNOFF_CMM : DInt := 100000;   // Break downstream offset [mm/100]
      CONST_DBREAKUPOFF_CMM : DInt := 100000;   // Break upstream offset [mm/100]
   END_VAR
BEGIN

REGION Network 1: CPUs
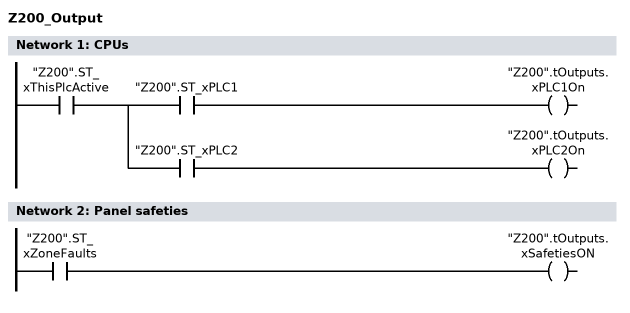
   RUNG wire#powerrail
      Contact( "Z200".ST_xThisPlcActive )
      wire#w1
      Contact( "Z200".ST_xPLC1 )
      Coil( "Z200".tOutputs.xPLC1On )
   END_RUNG
   RUNG wire#w1
      Contact( "Z200".ST_xPLC2 )
      Coil( "Z200".tOutputs.xPLC2On )
   END_RUNG
   // the same network as SCL:
   "Z200".tOutputs.xPLC1On := "Z200".ST_xThisPlcActive AND "Z200".ST_xPLC1;
   "Z200".tOutputs.xPLC2On := "Z200".ST_xThisPlcActive AND "Z200".ST_xPLC2;
END_REGION

REGION Network 2: Panel safeties
   RUNG wire#powerrail
      Contact( "Z200".ST_xZoneFaults )
      Coil( "Z200".tOutputs.xSafetiesON )
   END_RUNG
   // the same network as SCL:
   "Z200".tOutputs.xSafetiesON := "Z200".ST_xZoneFaults;
END_REGION
END_FUNCTION

// folder: 03_Programs_Logics/MCC1200/10_YCuts

FUNCTION_BLOCK "FB_YCuts_V1.00"   // FB9, LAD
TITLE = YCuts machine V1.00
{ S7_Optimized_Access := 'TRUE' }
VERSION : 0.1
   VAR_INPUT
      IN_dMachineIndex : DInt;   // Tracking machine index
      IN_dYCUTID : DInt;   // YCut identifier (0=M256A 1=M256B etc...)
      IN_dTrackNewCapIndex : DInt;   // New cap available on tracking index
      IN_xCycleON : Bool;   // Cycle ON
      IN_xGeneralReset : Bool;   // General reset
      IN_xResetAlarms : Bool;   // Reset alarms
      IN_xFaultsEnabled : Bool;   // Faults enabled
      IN_tID : Conn_Any;   // Connection ID
      IN_tIDeviceData : "UDT_YCut_IdeviceFromBridge";   // IDeviceData from bridge
      IN_xSimulationActive : Bool;   // Enable simulation (EXPERT USER)
      IN_dGlassBreakMachineIndex : DInt;   // Glass break machine index
   END_VAR
   VAR_OUTPUT
      OUT_tIDeviceData : "UDT_YCut_IdeviceToBridge";   // IDeviceData to bridge
      OUT_tBridgeStatus : Struct
         dBridgeStatus : DInt;   // Bridge actual status (1=OutOfProd 3=InProd 4=GlassBreak)
         rgxHeadProdOn : Array[0.."DMAXYHEADS_IND"] of Bool;   // Head#x production status
         rgxFireON : Array[0.."DMAXYHEADS_IND"] of Bool;   // Head#x fire status
         rgxArmON : Array[0.."DMAXYHEADS_IND"] of Bool;   // Head#x arm status
         rgdPosition_cmm : Array[0.."DMAXYHEADS_IND"] of DInt;   // Head#x position [mm/100]
      END_STRUCT;
   END_VAR
   VAR_IN_OUT
      INO_tTrack : "UDT_CapData_Tracking";   // Tracking plate
      INO_tEnc : "UDT_Encoder";   // Encoder data
      INO_tRibbon : "UDT_RibbonData";   // Ribbon data
   END_VAR
   VAR RETAIN
      tHMW : Struct   // HMI Write data
         xUpdateDistSnap : Bool;   // Update distance from snap roll {x|x|x|x|M}
         dDistanceFromSnaproll_cmm : DInt;   // Distance from snaproll [mm/100] [mm/100] {mm/100|mm|0|60000|M}
      END_STRUCT;
      tHMR : Struct   // HMI Read data
         dDistanceFromSnaproll_cmm : DInt;   // Distance from snaproll [mm/100] {mm/100|mm|0|60000|M}
      END_STRUCT;
   END_VAR
   VAR
      tALM : Struct   // HMI Alarms
         tS : Struct   // Stopping faults
            xTOutSendData : Bool;   // Timeout send data to bridge
            xSpare_1 : Bool;
            xSpare_2 : Bool;
            xSpare_3 : Bool;
            xSpare_4 : Bool;
            xSpare_5 : Bool;
            xSpare_6 : Bool;
            xSpare_7 : Bool;
            xSpare_8 : Bool;
            xSpare_9 : Bool;
            xSpare_10 : Bool;
            xSpare_11 : Bool;
            xSpare_12 : Bool;
            xSpare_13 : Bool;
            xSpare_14 : Bool;
            xSpare_15 : Bool;
            xSpare_16 : Bool;
            xSpare_17 : Bool;
            xSpare_18 : Bool;
            xSpare_19 : Bool;
            xSpare_20 : Bool;
            xSpare_21 : Bool;
            xSpare_22 : Bool;
            xSpare_23 : Bool;
            xSpare_24 : Bool;
            xSpare_25 : Bool;
            xSpare_26 : Bool;
            xSpare_27 : Bool;
            xSpare_28 : Bool;
            xSpare_29 : Bool;
            xSpare_30 : Bool;
            xSpare_31 : Bool;
         END_STRUCT;
         tF : Struct   // Faults
            xSpare_0 : Bool;
            xSpare_1 : Bool;
            xSpare_2 : Bool;
            xSpare_3 : Bool;
            xSpare_4 : Bool;
            xSpare_5 : Bool;
            xSpare_6 : Bool;
            xSpare_7 : Bool;
            xSpare_8 : Bool;
            xSpare_9 : Bool;
            xSpare_10 : Bool;
            xSpare_11 : Bool;
            xSpare_12 : Bool;
            xSpare_13 : Bool;
            xSpare_14 : Bool;
            xSpare_15 : Bool;
            xSpare_16 : Bool;
            xSpare_17 : Bool;
            xSpare_18 : Bool;
            xSpare_19 : Bool;
            xSpare_20 : Bool;
            xSpare_21 : Bool;
            xSpare_22 : Bool;
            xSpare_23 : Bool;
            xSpare_24 : Bool;
            xSpare_25 : Bool;
            xSpare_26 : Bool;
            xSpare_27 : Bool;
            xSpare_28 : Bool;
            xSpare_29 : Bool;
            xSpare_30 : Bool;
            xSpare_31 : Bool;
         END_STRUCT;
         tW : Struct   // Warnings
            xSpare_0 : Bool;
            xSpare_1 : Bool;
            xSpare_2 : Bool;
            xSpare_3 : Bool;
            xSpare_4 : Bool;
            xSpare_5 : Bool;
            xSpare_6 : Bool;
            xSpare_7 : Bool;
            xSpare_8 : Bool;
            xSpare_9 : Bool;
            xSpare_10 : Bool;
            xSpare_11 : Bool;
            xSpare_12 : Bool;
            xSpare_13 : Bool;
            xSpare_14 : Bool;
            xSpare_15 : Bool;
            xSpare_16 : Bool;
            xSpare_17 : Bool;
            xSpare_18 : Bool;
            xSpare_19 : Bool;
            xSpare_20 : Bool;
            xSpare_21 : Bool;
            xSpare_22 : Bool;
            xSpare_23 : Bool;
            xSpare_24 : Bool;
            xSpare_25 : Bool;
            xSpare_26 : Bool;
            xSpare_27 : Bool;
            xSpare_28 : Bool;
            xSpare_29 : Bool;
            xSpare_30 : Bool;
            xSpare_31 : Bool;
         END_STRUCT;
      END_STRUCT;
      ST_xPhaseInProgress : Bool;   // Phases are in progress
      ST_xPhaseInProgressNetwork : Bool;   // Phase are in progress network
      AUX_xValidUpCap : Bool;   // Upstream cap is valid
      AUX_xValidDwCap : Bool;   // Downstream cap is valid
      AUX_dUpCapIndex : DInt;   // Index of the upstream cap
      AUX_dDwCapIndex : DInt;   // Index of the downstream cap
      OS_xNewCapUp : Bool;   // New cap arrived upstream
      OS_xNewCapDw : Bool;   // New cap arrived downstream
      OS_xNewCap : Bool;   // New cap arrived
      ST_xStoppingFaults : Bool;   // Stopping faults
      ST_xFaults : Bool;   // Faults
      ST_xWarnings : Bool;   // Warnings
      ST_xOutputEnabled : Bool;   // Output enabled
      ST_xGlassBreak : Bool;   // Glass break under bridge
      AUX_xUpIsQuality : Bool;   // Upstream cap is a quality cap
      AUX_xDwIsQuality : Bool;   // Downstream cap is a quality cap
      tPhases : Struct   // Phases
         xPlateUnderBridge : Bool;   // Plate in passage under bridge
         xSpare1 : Bool;
         xSpare2 : Bool;
         xSpare3 : Bool;
         xSpare4 : Bool;
         xSpare5 : Bool;
         xSpare6 : Bool;
         xSpare7 : Bool;
         xSpare8 : Bool;
         xSpare9 : Bool;
         xSpare10 : Bool;
         xSpare11 : Bool;
         xSpare12 : Bool;
         xSpare13 : Bool;
         xSpare14 : Bool;
         xSpare15 : Bool;
         xSpare16 : Bool;
         xSpare17 : Bool;
         xSpare18 : Bool;
         xSpare19 : Bool;
         xSpare20 : Bool;
         xSpare21 : Bool;
         xSpare22 : Bool;
         xSpare23 : Bool;
         xSpare24 : Bool;
         xSpare25 : Bool;
         xSpare26 : Bool;
         xSpare27 : Bool;
         xSpare28 : Bool;
         xSpare29 : Bool;
         xSpare30 : Bool;
         xSpare31 : Bool;
      END_STRUCT;
      tPhasesNetwork : Struct
         xSendMissionInProgr : Bool;   // Send mission data in progress
         xEndSendMissionInProgr : Bool;   // End send mission in progress
         xSendSyncroInProgr : Bool;   // Send syncro in progress
         xEndSendSyncroInProgr : Bool;   // End send syncro in progress
         xSpare4 : Bool;
         xSpare5 : Bool;
         xSpare6 : Bool;
         xSpare7 : Bool;
         xSpare8 : Bool;
         xSpare9 : Bool;
         xSpare10 : Bool;
         xSpare11 : Bool;
         xSpare12 : Bool;
         xSpare13 : Bool;
         xSpare14 : Bool;
         xSpare15 : Bool;
         xSpare16 : Bool;
         xSpare17 : Bool;
         xSpare18 : Bool;
         xSpare19 : Bool;
         xSpare20 : Bool;
         xSpare21 : Bool;
         xSpare22 : Bool;
         xSpare23 : Bool;
         xSpare24 : Bool;
         xSpare25 : Bool;
         xSpare26 : Bool;
         xSpare27 : Bool;
         xSpare28 : Bool;
         xSpare29 : Bool;
         xSpare30 : Bool;
         xSpare31 : Bool;
      END_STRUCT;
      FB_BSEND : BSEND;   // BSend instance
      AUX_tSendDataToBridge : Struct   // Send data to bridge
         tSyncroData : Struct
            dMissionID : DInt;
            dSynchroValue_cmm : DInt;
            dSpare : Array[0..7] of DInt;
            xSpare : Array[0..15] of Bool;
            dSpare2 : Array[0..2] of DInt;
            iSpare : Int;
         END_STRUCT;
         tMissionData : Struct
            dMissionID : DInt;
            dMissionStart_cmm : DInt;
            dMissionEnd_cmm : DInt;
            dTrackingDbNumber : DInt;
            dSpare1 : Array[0..9] of DInt;
            rgxFireRequest : Array[0..31] of Bool;
            rgdHeadsPosition_cmm : Array[0..15] of DInt;
            dSpare2 : Array[0..14] of DInt;
         END_STRUCT;
      END_STRUCT;
      ST_xRetrySendMission : Bool;   // Retry send mission
      ST_xRetrySendSyncro : Bool;   // Retry send syncro
      AUX_xCheckPlateCutDone : Bool;   // Check the plate for cut done analysis
      AUX_dActualRecoverWander_cmm : DInt;   // Actual recovered wander [mm/100]
      AUX_xQualityCap : Bool;   // Plate in passage is quality cap
   END_VAR
   VAR_TEMP
      TMP_dwValue : DWord;
      TMP_xCompileMissionData : Bool;
      TMP_dIndex : DInt;
      TMP_wPackLength : Word;
      TMP_xRetrySendMissionWithNewMission : Bool;
      TMP_xRetrySendSyncroWithNewSyncro : Bool;
      TMP_xCompileSyncroData : Bool;
      TMP_xNewCapAvailable : Bool;
      TMP_wValue : Word;
      TMP_dPercLength_cmm : DInt;
      TMP_dOpenGatePosition_cmm : DInt;
      TMP_dCloseGatePosition_cmm : DInt;
      TMP_dEncOnYCut_cmm : DInt;
      TMP_dValue_cmm : DInt;
      TMP_xRequestIsNotDone : Bool;
      TMP_xTripleEdgeSituation : Bool;
      TMP_dOppositeBridgeIndex : DInt;
   END_VAR
   VAR CONSTANT
      CONST_DBREAKDOWNOFF_CMM : DInt := 50000;   // Break downstream offset [mm/100]
      CONST_DBREAKUPOFF_CMM : DInt := 50000;   // Break upstream offset [mm/100]
      CONST_TRIPLE_FIRSTHEAD : DInt := 0;   // Triple edge first head
      CONST_TRIPLE_LASTHEAD : DInt := 8;   // Triple edge last head
   END_VAR
BEGIN

REGION Network 1: ####_CONSTANTS_####
END_REGION

REGION Network 2: ####_MATCH_####
END_REGION

REGION Network 3 (SCL): General reset clean
   IF #IN_xGeneralReset THEN

       #TMP_dwValue := 0;

       SCATTER(IN:=#TMP_dwValue,
               OUT=>#tPhases);

       SCATTER(IN:=#TMP_dwValue,
               OUT=>#tPhasesNetwork);


   END_IF;
END_REGION

REGION Network 4 (SCL): Move data information to tracking
   #INO_tTrack.rgtTrackMachine[#IN_dMachineIndex].tUserData.dSetDistanceSnap_cmm := #tHMR.dDistanceFromSnaproll_cmm;
   #INO_tTrack.rgtTrackMachine[#IN_dMachineIndex].tUserData.dSetMachReacTime_ms := 0;
END_REGION

REGION Network 5 (SCL): Manage tracking call

   #OS_xNewCapUp := FALSE;
   #OS_xNewCapDw := FALSE;
   #OS_xNewCap := FALSE;

   IF #INO_tTrack.rgtTrackMachine[#IN_dMachineIndex].tUserData.xGetPosReach THEN

       #OS_xNewCap := TRUE;

       IF #INO_tTrack.rgtTrackMachine[#IN_dMachineIndex].tUserData.dGetUpstremIndex >= 0 THEN
           #AUX_xValidUpCap := TRUE;
           #OS_xNewCapUp := TRUE;            
           #AUX_dUpCapIndex := #INO_tTrack.rgtTrackMachine[#IN_dMachineIndex].tUserData.dGetUpstremIndex;
       ELSE
           #AUX_xValidUpCap := FALSE;
           #OS_xNewCapUp := FALSE;            
           #AUX_dUpCapIndex := 0;
       END_IF;

